REGION Network 4: Управление запуском
   RUNG wire#powerrail
      Contact( #Data )
      I_Contact( #Inverse )
      wire#w1
      I_Contact( #Hand )
      wire#w2
      S_SR(operand := #Start_M, r1 := wire#w4)
      Coil( #Signal )
   END_RUNG
   RUNG wire#powerrail
      I_Contact( #Data )
      Contact( #Inverse )
   END_RUNG wire#w1
   RUNG wire#powerrail
      Contact( #Hand )
      Contact( #Start_M )
   END_RUNG wire#w2
   RUNG wire#powerrail
      Contact( #Data )
      Contact( #Inverse )
      wire#w3
      I_Contact( #Hand )
   END_RUNG wire#w4
   RUNG wire#powerrail
      I_Contact( #Data )
      I_Contact( #Inverse )
   END_RUNG wire#w3
   RUNG wire#powerrail
      Contact( #Hand )
      I_Contact( #Start_M )
   END_RUNG wire#w4
   // the same network as SCL:
   #_w1 := (((#Data AND #Inverse) OR (NOT #Data AND NOT #Inverse)) AND NOT #Hand) OR (#Hand AND NOT #Start_M);
   IF (((#Data AND NOT #Inverse) OR (NOT #Data AND #Inverse)) AND NOT #Hand) OR (#Hand AND #Start_M) THEN
       #Start_M := TRUE;   // SR flip-flop
   END_IF;
   IF #_w1 THEN #Start_M := FALSE; END_IF;
   #Signal := #Start_M;
END_REGION

REGION Network 5: Блок таймеров
   RUNG wire#powerrail
      "Time_s"(pulse := #pulse, T := #Filter_On)
      "Time_s"(pulse := #pulse, T := #Filter_Off)
   END_RUNG
   // the same network as SCL:
   "Time_s"(pulse := #pulse, T := #Filter_On, ENO => #_w1);
   IF #_w1 THEN "Time_s"(pulse := #pulse, T := #Filter_Off); END_IF;
END_REGION
END_FUNCTION_BLOCK

FUNCTION_BLOCK "DO_ex"   // FB101, LAD
{ S7_Optimized_Access := 'FALSE' }
VERSION : 0.1
   VAR_IN_OUT
      Start_A : Bool;   // Управляющий сигнал из программы
      pulse : Bool;   // Частота длительности импульса
      Q : Bool;   // Выходной сигнал контроллера
   END_VAR
   VAR
      Hand : Bool;   // 0 - Авто, 1 - Ручной
      Start_M : Bool;   // Запуск в ручном режиме
      Simulation : Bool;   // Режим симуляции
      Inverse : Bool;   // Инверсия выхода
      Impulse : Bool;   // Импульсный режим
      T_Impulse : Struct   // Длительность импульса
         SP : Int := 5;
         Now : Int;
         "Exit" : Bool;
         Start : Bool;
         Pause : Bool;
         Reset : Bool;
      END_STRUCT;
   END_VAR
   VAR_TEMP   // added for the SCL form of the ladder/FBD networks
      _w1 : Bool;
   END_VAR
BEGIN

REGION Network 1: Устройство в ручном режиме
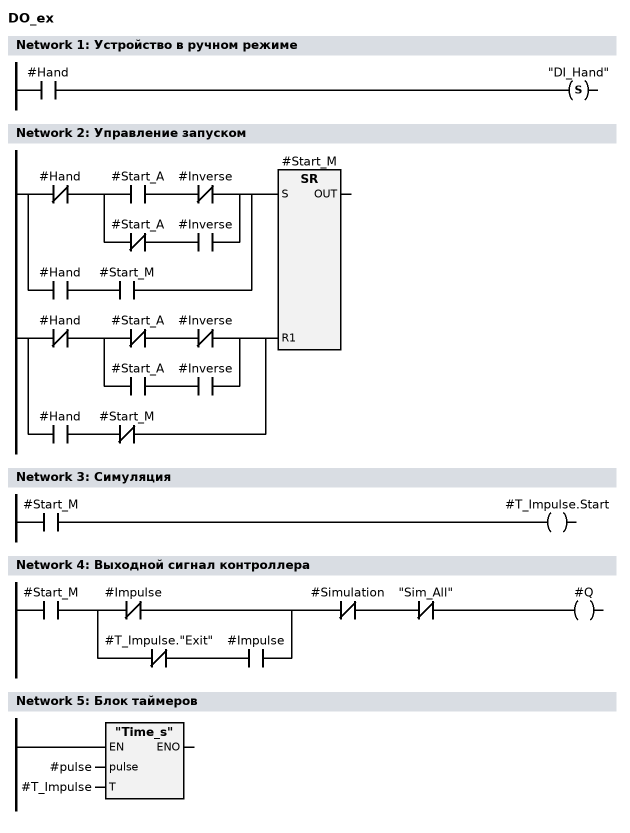
   RUNG wire#powerrail
      Contact( #Hand )
      S_Coil( "DI_Hand" )
   END_RUNG
   // the same network as SCL:
   IF #Hand THEN "DI_Hand" := TRUE; END_IF;
END_REGION

REGION Network 2: Управление запуском
   RUNG wire#powerrail
      I_Contact( #Hand )
      wire#w1
      Contact( #Start_A )
      I_Contact( #Inverse )
      wire#w2
      S_SR(operand := #Start_M, r1 := wire#w4)
   END_RUNG
   RUNG wire#w1
      I_Contact( #Start_A )
      Contact( #Inverse )
   END_RUNG wire#w2
   RUNG wire#powerrail
      Contact( #Hand )
      Contact( #Start_M )
   END_RUNG wire#w2
   RUNG wire#powerrail
      I_Contact( #Hand )
      wire#w3
      I_Contact( #Start_A )
      I_Contact( #Inverse )
   END_RUNG wire#w4
   RUNG wire#w3
      Contact( #Start_A )
      Contact( #Inverse )
   END_RUNG wire#w4
   RUNG wire#powerrail
      Contact( #Hand )
      I_Contact( #Start_M )
   END_RUNG wire#w4
   // the same network as SCL:
   #_w1 := (NOT #Hand AND ((NOT #Start_A AND NOT #Inverse) OR (#Start_A AND #Inverse))) OR (#Hand AND NOT #Start_M);
   IF (NOT #Hand AND ((#Start_A AND NOT #Inverse) OR (NOT #Start_A AND #Inverse))) OR (#Hand AND #Start_M) THEN
       #Start_M := TRUE;   // SR flip-flop
   END_IF;
   IF #_w1 THEN #Start_M := FALSE; END_IF;
END_REGION

REGION Network 3: Симуляция
   RUNG wire#powerrail
      Contact( #Start_M )
      Coil( #T_Impulse.Start )
   END_RUNG
   // the same network as SCL:
   #T_Impulse.Start := #Start_M;
END_REGION

REGION Network 4: Выходной сигнал контроллера
   RUNG wire#powerrail
      Contact( #Start_M )
      wire#w1
      I_Contact( #Impulse )
      wire#w2
      I_Contact( #Simulation )
      I_Contact( "Sim_All" )
      Coil( #Q )
   END_RUNG
   RUNG wire#w1
      I_Contact( #T_Impulse."Exit" )
      Contact( #Impulse )
   END_RUNG wire#w2
   // the same network as SCL:
   #Q := #Start_M AND (NOT #Impulse OR (NOT #T_Impulse."Exit" AND #Impulse)) AND NOT #Simulation AND NOT "Sim_All";
END_REGION

REGION Network 5: Блок таймеров
   RUNG wire#powerrail
      "Time_s"(pulse := #pulse, T := #T_Impulse)
   END_RUNG
   // the same network as SCL:
   "Time_s"(pulse := #pulse, T := #T_Impulse);
END_REGION
END_FUNCTION_BLOCK

FUNCTION_BLOCK "DRV_Micro"   // FB104, LAD
{ S7_Optimized_Access := 'FALSE' }
VERSION : 0.1
   VAR_INPUT
      Start_A : Bool;   // Запрос запуска
      FB : Bool;   // ОС
      Reset : Bool;   // Сброс аварий
      All_Block : Bool;   // Блокировка
   END_VAR
   VAR_OUTPUT
      CMD : Bool;   // Команда
   END_VAR
   VAR_IN_OUT
      Alarm : Bool;   // Авария
   END_VAR
   VAR
      Hand : Bool;   // Ручной режим
      Start_M : Bool;   // Запуск в ручном режиме
      No_FB : Bool;   // Не использовать ОС
      ON : Bool;   // Успешно запущено
      OFF : Bool;   // Успешно остановлено
      Status : Int;   // Статус устройства / Статус привода
      Wait_On : Struct   // Ожидание ОС контактора / Время на запуск
         SP : Int := 2;
         Now : Int;
         "Exit" : Bool;
         Start : Bool;
         Pause : Bool;
         Reset : Bool;
      END_STRUCT;
      Wait_Off : Struct   // Ожидание концевиков / Время на останов
         SP : Int := 2;
         Now : Int;
         "Exit" : Bool;
         Start : Bool;
         Pause : Bool;
         Reset : Bool;
      END_STRUCT;
   END_VAR
   VAR_TEMP   // added for the SCL form of the ladder/FBD networks
      _w1 : Bool;
      _w2 : Bool;
   END_VAR
BEGIN

REGION Network 1: Управление запуском / дискретный управляющий сигнал
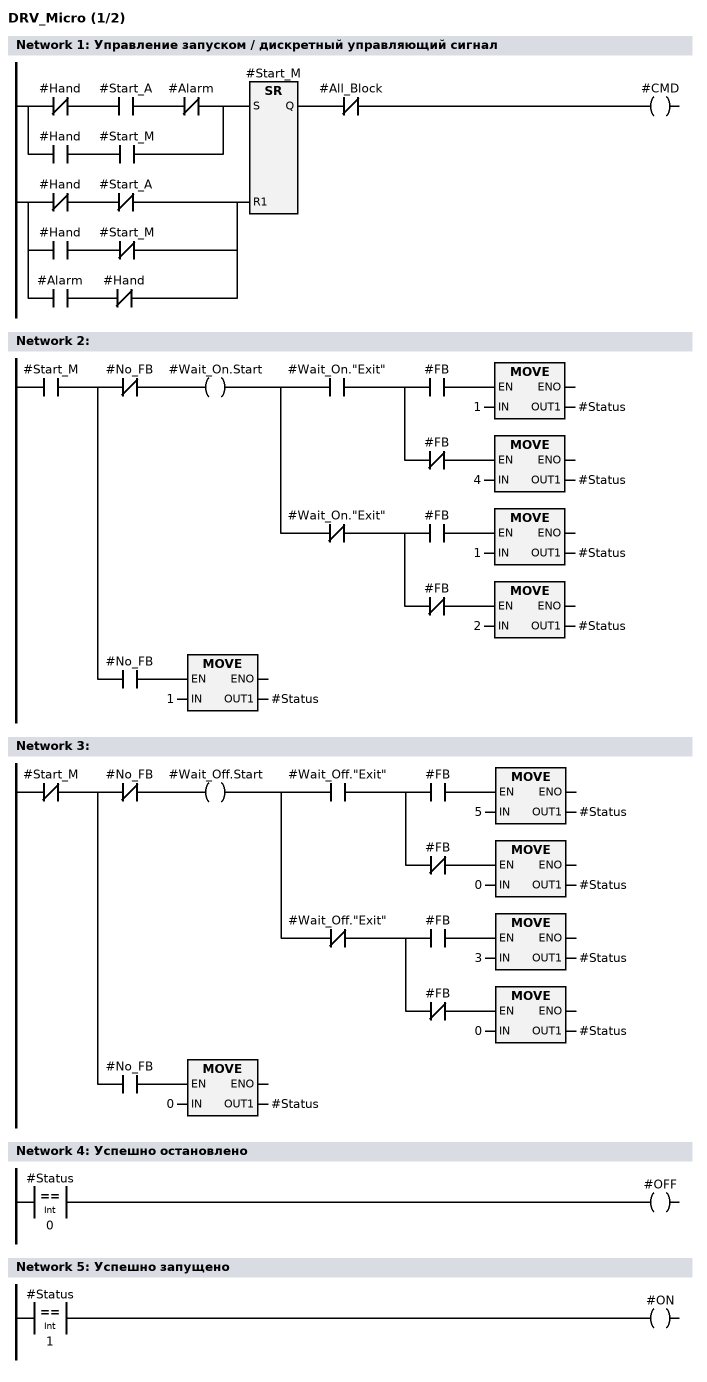
   RUNG wire#powerrail
      I_Contact( #Hand )
      Contact( #Start_A )
      I_Contact( #Alarm )
      wire#w1
      S_SR(operand := #Start_M, r1 := wire#w2)
      I_Contact( #All_Block )
      Coil( #CMD )
   END_RUNG
   RUNG wire#powerrail
      Contact( #Hand )
      Contact( #Start_M )
   END_RUNG wire#w1
   RUNG wire#powerrail
      I_Contact( #Hand )
      I_Contact( #Start_A )
   END_RUNG wire#w2
   RUNG wire#powerrail
      Contact( #Hand )
      I_Contact( #Start_M )
   END_RUNG wire#w2
   RUNG wire#powerrail
      Contact( #Alarm )
      I_Contact( #Hand )
   END_RUNG wire#w2
   // the same network as SCL:
   #_w1 := (NOT #Hand AND NOT #Start_A) OR (#Hand AND NOT #Start_M) OR (#Alarm AND NOT #Hand);
   IF (NOT #Hand AND #Start_A AND NOT #Alarm) OR (#Hand AND #Start_M) THEN
       #Start_M := TRUE;   // SR flip-flop
   END_IF;
   IF #_w1 THEN #Start_M := FALSE; END_IF;
   #CMD := #Start_M AND NOT #All_Block;
END_REGION

REGION Network 2
   RUNG wire#powerrail
      Contact( #Start_M )
      wire#w1
      I_Contact( #No_FB )
      Coil( #Wait_On.Start )
      wire#w2
      Contact( #Wait_On."Exit" )
      wire#w3
      Contact( #FB )
      Move(in := 1, out1 => #Status)
   END_RUNG
   RUNG wire#w3
      I_Contact( #FB )
      Move(in := 4, out1 => #Status)
   END_RUNG
   RUNG wire#w2
      I_Contact( #Wait_On."Exit" )
      wire#w4
      Contact( #FB )
      Move(in := 1, out1 => #Status)
   END_RUNG
   RUNG wire#w4
      I_Contact( #FB )
      Move(in := 2, out1 => #Status)
   END_RUNG
   RUNG wire#w1
      Contact( #No_FB )
      Move(in := 1, out1 => #Status)
   END_RUNG
   // the same network as SCL:
   #Wait_On.Start := #Start_M AND NOT #No_FB;
   #_w1 := #Wait_On.Start AND #Wait_On."Exit";
   IF #_w1 AND #FB THEN #Status := 1; END_IF;
   IF #_w1 AND NOT #FB THEN #Status := 4; END_IF;
   #_w2 := #Wait_On.Start AND NOT #Wait_On."Exit";
   IF #_w2 AND #FB THEN #Status := 1; END_IF;
   IF #_w2 AND NOT #FB THEN #Status := 2; END_IF;
   IF #Start_M AND #No_FB THEN #Status := 1; END_IF;
END_REGION

REGION Network 3
   RUNG wire#powerrail
      I_Contact( #Start_M )
      wire#w1
      I_Contact( #No_FB )
      Coil( #Wait_Off.Start )
      wire#w2
      Contact( #Wait_Off."Exit" )
      wire#w3
      Contact( #FB )
      Move(in := 5, out1 => #Status)
   END_RUNG
   RUNG wire#w3
      I_Contact( #FB )
      Move(in := 0, out1 => #Status)
   END_RUNG
   RUNG wire#w2
      I_Contact( #Wait_Off."Exit" )
      wire#w4
      Contact( #FB )
      Move(in := 3, out1 => #Status)
   END_RUNG
   RUNG wire#w4
      I_Contact( #FB )
      Move(in := 0, out1 => #Status)
   END_RUNG
   RUNG wire#w1
      Contact( #No_FB )
      Move(in := 0, out1 => #Status)
   END_RUNG
   // the same network as SCL:
   #Wait_Off.Start := NOT #Start_M AND NOT #No_FB;
   #_w1 := #Wait_Off.Start AND #Wait_Off."Exit";
   IF #_w1 AND #FB THEN #Status := 5; END_IF;
   IF #_w1 AND NOT #FB THEN #Status := 0; END_IF;
   #_w2 := #Wait_Off.Start AND NOT #Wait_Off."Exit";
   IF #_w2 AND #FB THEN #Status := 3; END_IF;
   IF #_w2 AND NOT #FB THEN #Status := 0; END_IF;
   IF NOT #Start_M AND #No_FB THEN #Status := 0; END_IF;
END_REGION

REGION Network 4: Успешно остановлено
   RUNG wire#powerrail
      { S7_Templates := "SrcType := Int" } EQ_Contact(in1 := #Status, in2 := 0)
      Coil( #OFF )
   END_RUNG
   // the same network as SCL:
   #OFF := #Status = 0;
END_REGION

REGION Network 5: Успешно запущено
   RUNG wire#powerrail
      { S7_Templates := "SrcType := Int" } EQ_Contact(in1 := #Status, in2 := 1)
      Coil( #ON )
   END_RUNG
   // the same network as SCL:
   #ON := #Status = 1;
END_REGION

REGION Network 6: Авария
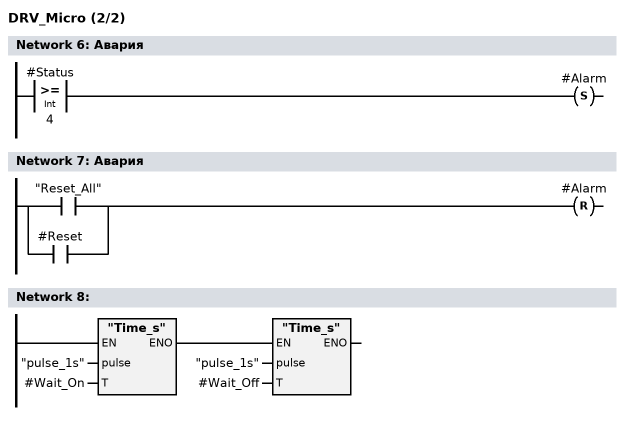
   RUNG wire#powerrail
      { S7_Templates := "SrcType := Int" } GE_Contact(in1 := #Status, in2 := 4)
      S_Coil( #Alarm )
   END_RUNG
   // the same network as SCL:
   IF #Status >= 4 THEN #Alarm := TRUE; END_IF;
END_REGION

REGION Network 7: Авария
   RUNG wire#powerrail
      Contact( "Reset_All" )
      wire#w1
      R_Coil( #Alarm )
   END_RUNG
   RUNG wire#powerrail
      Contact( #Reset )
   END_RUNG wire#w1
   // the same network as SCL:
   IF "Reset_All" OR #Reset THEN #Alarm := FALSE; END_IF;
END_REGION

REGION Network 8
   RUNG wire#powerrail
      "Time_s"(pulse := "pulse_1s", T := #Wait_On)
      "Time_s"(pulse := "pulse_1s", T := #Wait_Off)
   END_RUNG
   // the same network as SCL:
   "Time_s"(pulse := "pulse_1s", T := #Wait_On, ENO => #_w1);
   IF #_w1 THEN "Time_s"(pulse := "pulse_1s", T := #Wait_Off); END_IF;
END_REGION
END_FUNCTION_BLOCK

// folder: Modules

FUNCTION_BLOCK "DIx"   // FB200, LAD
{ S7_Optimized_Access := 'FALSE' }
VERSION : 0.1
// Input - входной сигнал контроллера
// pulse - частота фильтрации дребезга
// Signal - обработанный и отфильтрованный сигнал, используемый в дальнейшем
   VAR
      M1_FB_Ready : "DI_ex";   // I 0.0 - Мешалка 1 - готовность
      M1_FB_Run : "DI_ex";   // I 0.1 - Мешалка 1 - работа
      M2_FB_Ready : "DI_ex";   // I 0.2 - Мешалка 2 - готовность
      M2_FB_Run : "DI_ex";   // I 0.3 - Мешалка 2 - работа
      M3_FB_Ready : "DI_ex";   // I 0.4 - Мешалка 3 - готовность
      M3_FB_Run : "DI_ex";   // I 0.5 - Мешалка 3 - работа
      DD_FB_Ready : "DI_ex";   // I 0.6 - Дозатор сухого вещества - готовность
      Dos_FB_Run : "DI_ex";   // I 0.7 - Дозатор - работа
      DD_LLS : "DI_ex";   // I 1.0 - Дозатор сухого вещества - низкий уровень
      Vibro_FB_Ready : "DI_ex";   // I 1.1 - Вибратор - готовность
      Transporter : "DI_ex";   // I 1.2 - Пневмотранспортёр - готовность
      DL_FB_Ready : "DI_ex";   // I 1.3 - Дозатор жидкого вещества - готовность
      Dry_Run : "DI_ex";   // I 1.4 - Датчик протока
      AllBlock : "DI_ex";   // I 1.5 - Датчик перелива или Аварийная остановка
   END_VAR
   VAR_TEMP   // added for the SCL form of the ladder/FBD networks
      _w1 : Bool;
      _w2 : Bool;
   END_VAR
BEGIN

REGION Network 1: Мешалка 1
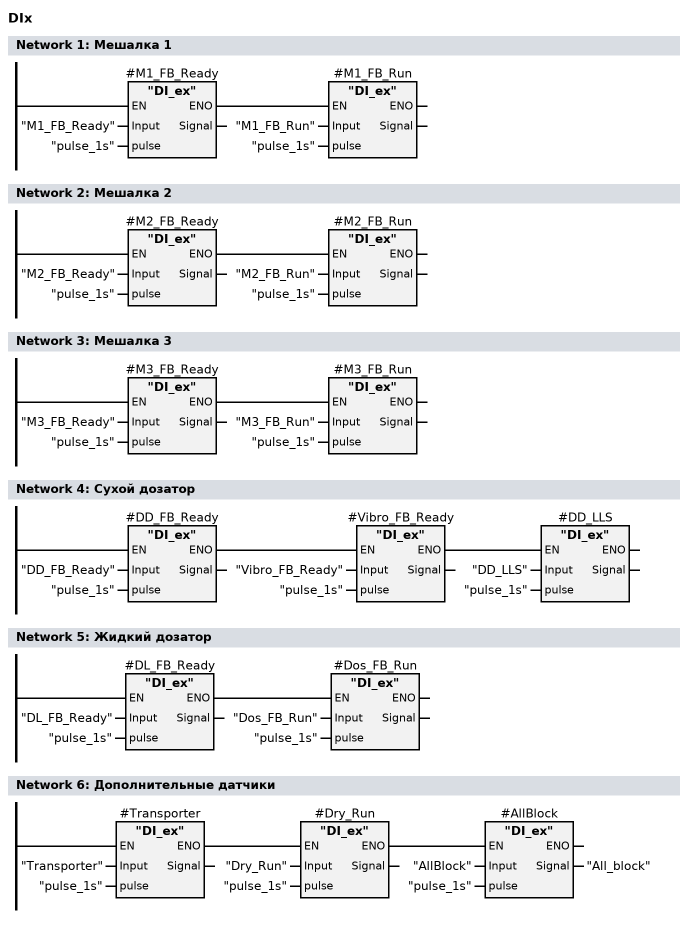
   RUNG wire#powerrail
      #M1_FB_Ready(Input := "M1_FB_Ready", pulse := "pulse_1s", Signal =>)
      #M1_FB_Run(Input := "M1_FB_Run", pulse := "pulse_1s", Signal =>)
   END_RUNG
   // the same network as SCL:
   #M1_FB_Ready(Input := "M1_FB_Ready", pulse := "pulse_1s", ENO => #_w1);   // "DI_ex"
   IF #_w1 THEN
       #M1_FB_Run(Input := "M1_FB_Run", pulse := "pulse_1s");   // "DI_ex"
   END_IF;
END_REGION

REGION Network 2: Мешалка 2
   RUNG wire#powerrail
      #M2_FB_Ready(Input := "M2_FB_Ready", pulse := "pulse_1s", Signal =>)
      #M2_FB_Run(Input := "M2_FB_Run", pulse := "pulse_1s", Signal =>)
   END_RUNG
   // the same network as SCL:
   #M2_FB_Ready(Input := "M2_FB_Ready", pulse := "pulse_1s", ENO => #_w1);   // "DI_ex"
   IF #_w1 THEN
       #M2_FB_Run(Input := "M2_FB_Run", pulse := "pulse_1s");   // "DI_ex"
   END_IF;
END_REGION

REGION Network 3: Мешалка 3
   RUNG wire#powerrail
      #M3_FB_Ready(Input := "M3_FB_Ready", pulse := "pulse_1s", Signal =>)
      #M3_FB_Run(Input := "M3_FB_Run", pulse := "pulse_1s", Signal =>)
   END_RUNG
   // the same network as SCL:
   #M3_FB_Ready(Input := "M3_FB_Ready", pulse := "pulse_1s", ENO => #_w1);   // "DI_ex"
   IF #_w1 THEN
       #M3_FB_Run(Input := "M3_FB_Run", pulse := "pulse_1s");   // "DI_ex"
   END_IF;
END_REGION

REGION Network 4: Сухой дозатор
   RUNG wire#powerrail
      #DD_FB_Ready(Input := "DD_FB_Ready", pulse := "pulse_1s", Signal =>)
      #Vibro_FB_Ready(Input := "Vibro_FB_Ready", pulse := "pulse_1s", Signal =>)
      #DD_LLS(Input := "DD_LLS", pulse := "pulse_1s", Signal =>)
   END_RUNG
   // the same network as SCL:
   #DD_FB_Ready(Input := "DD_FB_Ready", pulse := "pulse_1s", ENO => #_w1);   // "DI_ex"
   #Vibro_FB_Ready(EN := #_w1, Input := "Vibro_FB_Ready", pulse := "pulse_1s", ENO => #_w2);   // "DI_ex"
   IF #_w2 THEN
       #DD_LLS(Input := "DD_LLS", pulse := "pulse_1s");   // "DI_ex"
   END_IF;
END_REGION

REGION Network 5: Жидкий дозатор
   RUNG wire#powerrail
      #DL_FB_Ready(Input := "DL_FB_Ready", pulse := "pulse_1s", Signal =>)
      #Dos_FB_Run(Input := "Dos_FB_Run", pulse := "pulse_1s", Signal =>)
   END_RUNG
   // the same network as SCL:
   #DL_FB_Ready(Input := "DL_FB_Ready", pulse := "pulse_1s", ENO => #_w1);   // "DI_ex"
   IF #_w1 THEN
       #Dos_FB_Run(Input := "Dos_FB_Run", pulse := "pulse_1s");   // "DI_ex"
   END_IF;
END_REGION

REGION Network 6: Дополнительные датчики
   RUNG wire#powerrail
      #Transporter(Input := "Transporter", pulse := "pulse_1s", Signal =>)
      #Dry_Run(Input := "Dry_Run", pulse := "pulse_1s", Signal =>)
      #AllBlock(Input := "AllBlock", pulse := "pulse_1s", Signal => "All_block")
   END_RUNG
   // the same network as SCL:
   #Transporter(Input := "Transporter", pulse := "pulse_1s", ENO => #_w1);   // "DI_ex"
   #Dry_Run(EN := #_w1, Input := "Dry_Run", pulse := "pulse_1s", ENO => #_w2);   // "DI_ex"
   IF #_w2 THEN
       #AllBlock(Input := "AllBlock", pulse := "pulse_1s", Signal => "All_block");   // "DI_ex"
   END_IF;
END_REGION
END_FUNCTION_BLOCK

FUNCTION_BLOCK "DOx"   // FB201, LAD
{ S7_Optimized_Access := 'FALSE' }
VERSION : 0.1
// Start - управляющий сигнал из программы
// Q - выходной сигнал контроллера
// pulse - кратность времени в импульсном режиме
   VAR
      M1_CMD : "DO_ex";   // Q 0.0 - Мешалка 1 - запуск
      M2_CMD : "DO_ex";   // Q 0.1 - Мешалка 2 - запуск
      M3_CMD : "DO_ex";   // Q 0.2 - Мешалка 3 - запуск
      DD_CMD : "DO_ex";   // Q 0.3 - Дозатор сухого вещества - запуск
      Vibro_CMD : "DO_ex";   // Q 0.4 - Вибратор - запуск
      DL_CMD : "DO_ex";   // Q 0.5 - Дозатор жидкого вещества - запуск
      KC1_CMD : "DO_ex";   // Q 0.6 - Соленоидный клапан КС1
      LED_Dry_Run : "DO_ex";   // Q 0.7 - LED - сухой ход
      LED_Alarm : "DO_ex";   // Q 1.0 - LED - общая авария
      LED_Empty : "DO_ex";   // Q 1.1 - LED - бункер пуст
   END_VAR
   VAR_TEMP   // added for the SCL form of the ladder/FBD networks
      _w1 : Bool;
      _w2 : Bool;
   END_VAR
BEGIN

REGION Network 1: Мешалки 1-3
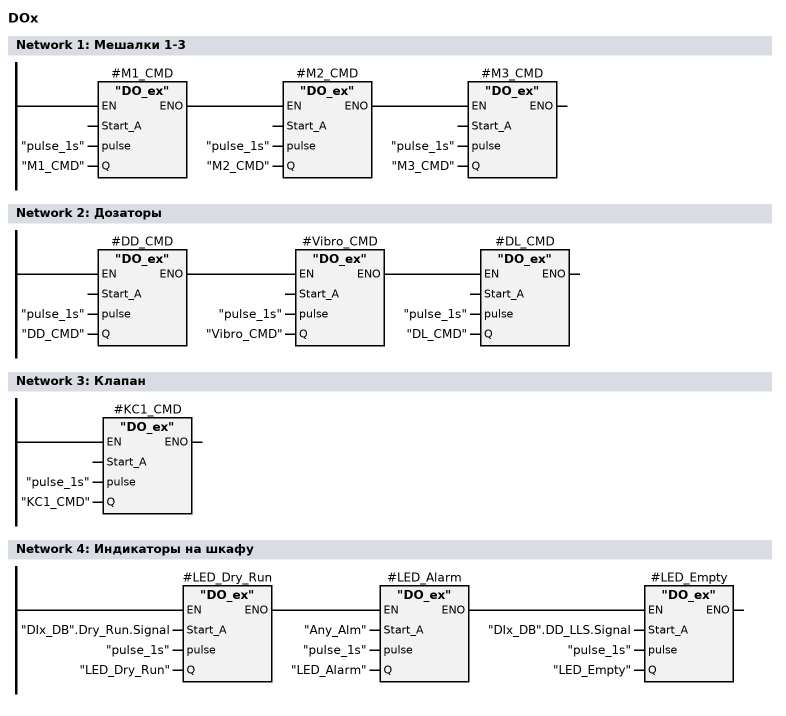
   RUNG wire#powerrail
      #M1_CMD(Start_A :=, pulse := "pulse_1s", Q := "M1_CMD")
      #M2_CMD(Start_A :=, pulse := "pulse_1s", Q := "M2_CMD")
      #M3_CMD(Start_A :=, pulse := "pulse_1s", Q := "M3_CMD")
   END_RUNG
   // the same network as SCL:
   #M1_CMD(pulse := "pulse_1s", Q := "M1_CMD", ENO => #_w1);   // "DO_ex"
   #M2_CMD(EN := #_w1, pulse := "pulse_1s", Q := "M2_CMD", ENO => #_w2);   // "DO_ex"
   IF #_w2 THEN
       #M3_CMD(pulse := "pulse_1s", Q := "M3_CMD");   // "DO_ex"
   END_IF;
END_REGION

REGION Network 2: Дозаторы
   RUNG wire#powerrail
      #DD_CMD(Start_A :=, pulse := "pulse_1s", Q := "DD_CMD")
      #Vibro_CMD(Start_A :=, pulse := "pulse_1s", Q := "Vibro_CMD")
      #DL_CMD(Start_A :=, pulse := "pulse_1s", Q := "DL_CMD")
   END_RUNG
   // the same network as SCL:
   #DD_CMD(pulse := "pulse_1s", Q := "DD_CMD", ENO => #_w1);   // "DO_ex"
   #Vibro_CMD(EN := #_w1, pulse := "pulse_1s", Q := "Vibro_CMD", ENO => #_w2);   // "DO_ex"
   IF #_w2 THEN
       #DL_CMD(pulse := "pulse_1s", Q := "DL_CMD");   // "DO_ex"
   END_IF;
END_REGION

REGION Network 3: Клапан
   RUNG wire#powerrail
      #KC1_CMD(Start_A :=, pulse := "pulse_1s", Q := "KC1_CMD")
   END_RUNG
   // the same network as SCL:
   #KC1_CMD(pulse := "pulse_1s", Q := "KC1_CMD");   // "DO_ex"
END_REGION

REGION Network 4: Индикаторы на шкафу
   RUNG wire#powerrail
      #LED_Dry_Run(Start_A := "DIx_DB".Dry_Run.Signal, pulse := "pulse_1s", Q := "LED_Dry_Run")
      #LED_Alarm(Start_A := "Any_Alm", pulse := "pulse_1s", Q := "LED_Alarm")
      #LED_Empty(Start_A := "DIx_DB".DD_LLS.Signal, pulse := "pulse_1s", Q := "LED_Empty")
   END_RUNG
   // the same network as SCL:
   #LED_Dry_Run(Start_A := "DIx_DB".Dry_Run.Signal, pulse := "pulse_1s", Q := "LED_Dry_Run", ENO => #_w1);   // "DO_ex"
   #LED_Alarm(EN := #_w1, Start_A := "Any_Alm", pulse := "pulse_1s", Q := "LED_Alarm", ENO => #_w2);   // "DO_ex"
   IF #_w2 THEN
       #LED_Empty(Start_A := "DIx_DB".DD_LLS.Signal, pulse := "pulse_1s", Q := "LED_Empty");   // "DO_ex"
   END_IF;
END_REGION
END_FUNCTION_BLOCK

FUNCTION_BLOCK "Micro"   // FB207, LAD
{ S7_Optimized_Access := 'FALSE' }
VERSION : 0.1
   VAR
      KC1 : "DRV_Micro";   // Соленоидный клапан
   END_VAR
   // KC1.No_FB := true;
BEGIN

REGION Network 1
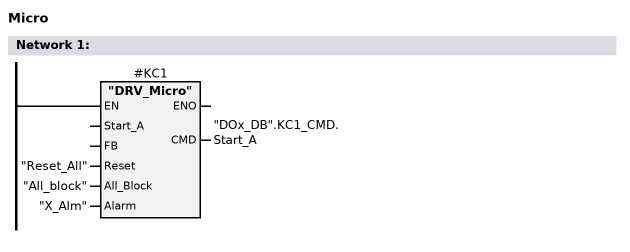
   RUNG wire#powerrail
      #KC1(Start_A :=, FB :=, Reset := "Reset_All", All_Block := "All_block", Alarm := "X_Alm", CMD => "DOx_DB".KC1_CMD.Start_A)
   END_RUNG
   // the same network as SCL:
   #KC1(Reset := "Reset_All", All_Block := "All_block", Alarm := "X_Alm", CMD => "DOx_DB".KC1_CMD.Start_A);   // "DRV_Micro"
END_REGION
END_FUNCTION_BLOCK

// folder: System

FUNCTION "DRV_pulse" : Void   // FC100, LAD
{ S7_Optimized_Access := 'FALSE' }
VERSION : 0.1
   VAR_TEMP   // added for the SCL form of the ladder/FBD networks
      _w1 : Bool;
      _w2 : Bool;
   END_VAR
BEGIN

REGION Network 1
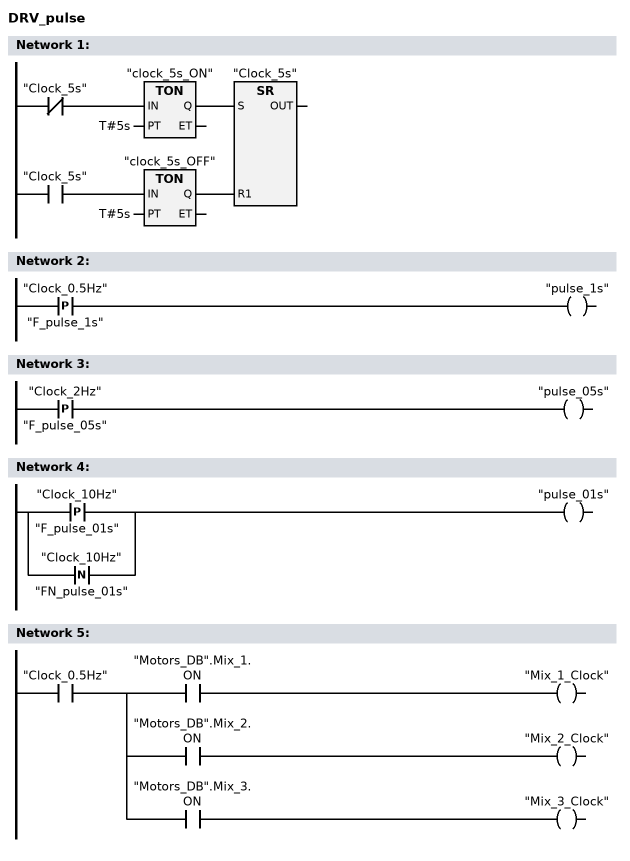
   "clock_5s_ON".TON(IN := NOT "Clock_5s", PT := T#5s);
   "clock_5s_OFF".TON(IN := "Clock_5s", PT := T#5s);
   IF "clock_5s_ON".Q THEN
       "Clock_5s" := TRUE;   // SR flip-flop
   END_IF;
   IF "clock_5s_OFF".Q THEN "Clock_5s" := FALSE; END_IF;
END_REGION

REGION Network 2
   RUNG wire#powerrail
      P_Contact(operand := "Clock_0.5Hz", bit := "F_pulse_1s")
      Coil( "pulse_1s" )
   END_RUNG
   // the same network as SCL:
   #_w1 := "Clock_0.5Hz" AND NOT "F_pulse_1s";   // rising edge of "Clock_0.5Hz"
   "F_pulse_1s" := "Clock_0.5Hz";
   "pulse_1s" := #_w1;
END_REGION

REGION Network 3
   RUNG wire#powerrail
      P_Contact(operand := "Clock_2Hz", bit := "F_pulse_05s")
      Coil( "pulse_05s" )
   END_RUNG
   // the same network as SCL:
   #_w1 := "Clock_2Hz" AND NOT "F_pulse_05s";   // rising edge of "Clock_2Hz"
   "F_pulse_05s" := "Clock_2Hz";
   "pulse_05s" := #_w1;
END_REGION

REGION Network 4
   RUNG wire#powerrail
      P_Contact(operand := "Clock_10Hz", bit := "F_pulse_01s")
      wire#w1
      Coil( "pulse_01s" )
   END_RUNG
   RUNG wire#powerrail
      N_Contact(operand := "Clock_10Hz", bit := "FN_pulse_01s")
   END_RUNG wire#w1
   // the same network as SCL:
   #_w1 := "Clock_10Hz" AND NOT "F_pulse_01s";   // rising edge of "Clock_10Hz"
   "F_pulse_01s" := "Clock_10Hz";
   #_w2 := NOT "Clock_10Hz" AND "FN_pulse_01s";   // falling edge of "Clock_10Hz"
   "FN_pulse_01s" := "Clock_10Hz";
   "pulse_01s" := #_w1 OR #_w2;
END_REGION

REGION Network 5
   RUNG wire#powerrail
      Contact( "Clock_0.5Hz" )
      wire#w1
      Contact( "Motors_DB".Mix_1.ON )
      Coil( "Mix_1_Clock" )
   END_RUNG
   RUNG wire#w1
      Contact( "Motors_DB".Mix_2.ON )
      Coil( "Mix_2_Clock" )
   END_RUNG
   RUNG wire#w1
      Contact( "Motors_DB".Mix_3.ON )
      Coil( "Mix_3_Clock" )
   END_RUNG
   // the same network as SCL:
   "Mix_1_Clock" := "Clock_0.5Hz" AND "Motors_DB".Mix_1.ON;
   "Mix_2_Clock" := "Clock_0.5Hz" AND "Motors_DB".Mix_2.ON;
   "Mix_3_Clock" := "Clock_0.5Hz" AND "Motors_DB".Mix_3.ON;
END_REGION
END_FUNCTION

FUNCTION "DRV_End" : Void   // FC101, LAD
{ S7_Optimized_Access := 'TRUE' }
VERSION : 0.1
BEGIN

REGION Network 1: Одно из устройств нижнего уровня в ручном режиме
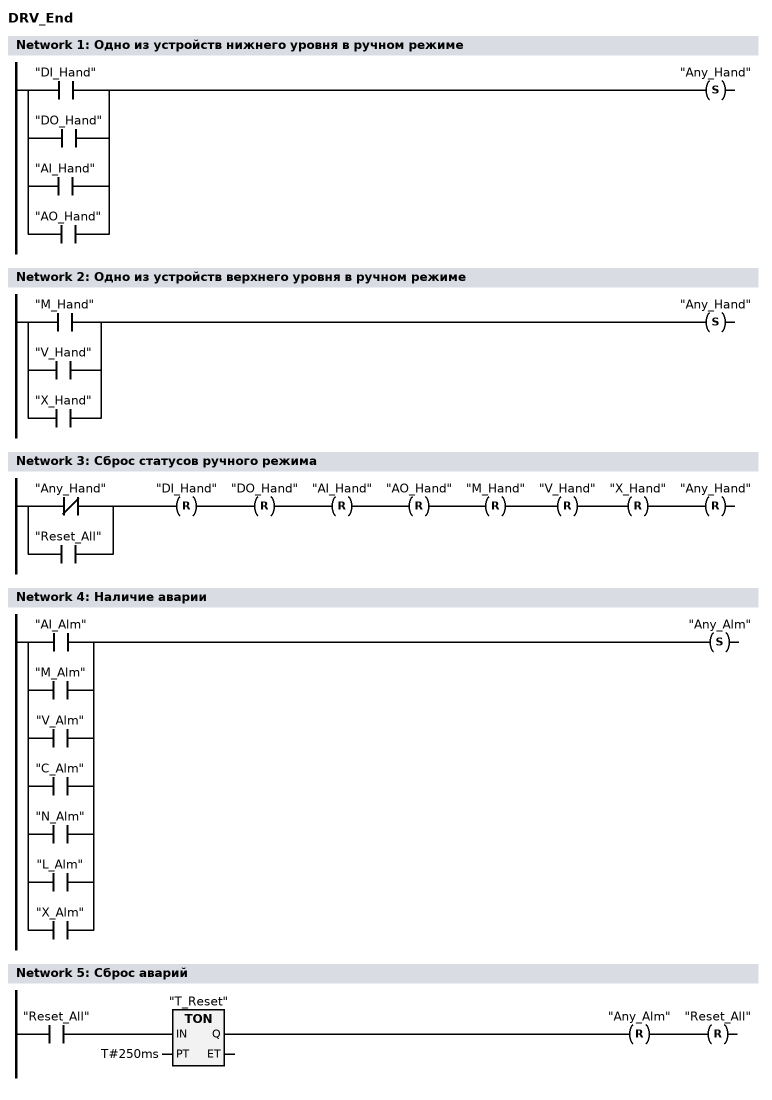
   RUNG wire#powerrail
      Contact( "DI_Hand" )
      wire#w1
      S_Coil( "Any_Hand" )
   END_RUNG
   RUNG wire#powerrail
      Contact( "DO_Hand" )
   END_RUNG wire#w1
   RUNG wire#powerrail
      Contact( "AI_Hand" )
   END_RUNG wire#w1
   RUNG wire#powerrail
      Contact( "AO_Hand" )
   END_RUNG wire#w1
   // the same network as SCL:
   IF "DI_Hand" OR "DO_Hand" OR "AI_Hand" OR "AO_Hand" THEN "Any_Hand" := TRUE; END_IF;
END_REGION

REGION Network 2: Одно из устройств верхнего уровня в ручном режиме
   RUNG wire#powerrail
      Contact( "M_Hand" )
      wire#w1
      S_Coil( "Any_Hand" )
   END_RUNG
   RUNG wire#powerrail
      Contact( "V_Hand" )
   END_RUNG wire#w1
   RUNG wire#powerrail
      Contact( "X_Hand" )
   END_RUNG wire#w1
   // the same network as SCL:
   IF "M_Hand" OR "V_Hand" OR "X_Hand" THEN "Any_Hand" := TRUE; END_IF;
END_REGION

REGION Network 3: Сброс статусов ручного режима
   RUNG wire#powerrail
      I_Contact( "Any_Hand" )
      wire#w1
      R_Coil( "DI_Hand" )
      R_Coil( "DO_Hand" )
      R_Coil( "AI_Hand" )
      R_Coil( "AO_Hand" )
      R_Coil( "M_Hand" )
      R_Coil( "V_Hand" )
      R_Coil( "X_Hand" )
      R_Coil( "Any_Hand" )
   END_RUNG
   RUNG wire#powerrail
      Contact( "Reset_All" )
   END_RUNG wire#w1
   // the same network as SCL:
   IF NOT "Any_Hand" OR "Reset_All" THEN
       "DI_Hand" := FALSE;
       "DO_Hand" := FALSE;
       "AI_Hand" := FALSE;
       "AO_Hand" := FALSE;
       "M_Hand" := FALSE;
       "V_Hand" := FALSE;
       "X_Hand" := FALSE;
       "Any_Hand" := FALSE;
   END_IF;
END_REGION

REGION Network 4: Наличие аварии
   RUNG wire#powerrail
      Contact( "AI_Alm" )
      wire#w1
      S_Coil( "Any_Alm" )
   END_RUNG
   RUNG wire#powerrail
      Contact( "M_Alm" )
   END_RUNG wire#w1
   RUNG wire#powerrail
      Contact( "V_Alm" )
   END_RUNG wire#w1
   RUNG wire#powerrail
      Contact( "C_Alm" )
   END_RUNG wire#w1
   RUNG wire#powerrail
      Contact( "N_Alm" )
   END_RUNG wire#w1
   RUNG wire#powerrail
      Contact( "L_Alm" )
   END_RUNG wire#w1
   RUNG wire#powerrail
      Contact( "X_Alm" )
   END_RUNG wire#w1
   // the same network as SCL:
   IF "AI_Alm" OR "M_Alm" OR "V_Alm" OR "C_Alm" OR "N_Alm" OR "L_Alm" OR "X_Alm" THEN
       "Any_Alm" := TRUE;
   END_IF;
END_REGION

REGION Network 5: Сброс аварий
   "T_Reset".TON(IN := "Reset_All", PT := T#250ms);
   IF "T_Reset".Q THEN
       "Any_Alm" := FALSE;
       "Reset_All" := FALSE;
   END_IF;
END_REGION
END_FUNCTION

FUNCTION "Converter" : Void   // FC102, LAD
TITLE = Драйвер линеаризации аналогового сигнала
{ S7_Optimized_Access := 'FALSE' }
VERSION : 0.1
   VAR_INPUT
      Converter : Struct
         Use_Min_In : Bool;   // Отсекать входные значения ниже минимума
         Use_Max_In : Bool;   // Отсекать входные значения выше максимума
         Use_Min_Out : Bool;   // Отсекать результат ниже минимума
         Use_Max_Out : Bool;   // Отсекать результат выше максимума
         Min_In : Real;   // Минимальный входной сигнал
         Max_In : Real;   // Максимальный входной сигнал
         Min_Out : Real;   // Минимальный выходной сигнал
         Max_Out : Real;   // Максимальный выходной сигнал
      END_STRUCT;
   END_VAR
   VAR_IN_OUT
      Signal : Real;   // Входной сигнал
      Result : Real;   // Результат линеаризации
   END_VAR
   VAR_TEMP
      Range_In : Real;   // Диапазон входного сигнала
      Range_Out : Real;   // Диапазон выходного сигнала
      T_T : Real;   // Соотношение диапазонов
      R_Sig : Real;   // Поправка на отрицательные значения
   END_VAR
BEGIN

REGION Network 1: Проверка нижнего уровня входного сигнала
